             // jog to position
             //*********************************************************************************************************
           ELSIF #tempJogToPosition THEN
             // set jog target position and configuration
             #instMC_MoveLinearAbsoute.Position[1] := #targetPosition.x;
             #instMC_MoveLinearAbsoute.Position[2] := #targetPosition.y;
             #instMC_MoveLinearAbsoute.Position[3] := #targetPosition.z;
             #instMC_MoveLinearAbsoute.Position[4] := #targetPosition.a;
             #instMC_MoveLinearAbsoute.CoordSystem := #coordSystem;
             #instMC_MoveLinearAbsoute.Velocity := #dynamics.path.velocity;
             #instMC_MoveLinearAbsoute.Acceleration := #dynamics.path.acceleration;
             #instMC_MoveLinearAbsoute.Deceleration := #dynamics.path.deceleration;
             #instMC_MoveLinearAbsoute.Jerk := #dynamics.path.jerk;
             #instMC_MoveLinearAbsoute.DynamicAdaption := #dynamics.dynamicAdaption;
           END_IF;

         END_REGION

         REGION STATE_TRANSITION

           // check if change of tool is required
           IF (#tool <> #statToolOld) THEN
             #statFBState := #FB_STATE_SET_TOOL;

             // check if orientation movement required
           ELSIF (((#jogDirection = 4) AND (#tempJogForward OR #tempJogBackward)) OR #tempJogToPosition)
             AND (#dynamics.orientation.velocity > 0.0 // check if change of orientation dynamics is required
             OR #dynamics.orientation.acceleration > 0.0
             OR #dynamics.orientation.deceleration > 0.0
             OR #dynamics.orientation.jerk > 0.0)
           THEN
             #statFBState := #FB_STATE_SET_DYNAMICS;

             // execute movement
           ELSE
             #statFBState := #FB_STATE_EXECUTE_MOVEMENT;
           END_IF;

         END_REGION

       #FB_STATE_SET_TOOL:

         REGION TOOL_CHANGE

           IF #axesGroup.StatusWord.%X6 // no motion command is acitve
             AND NOT #axesGroup.StatusWord.%X17 // not interrupted
             AND #axesGroup.StatusWord.%X12 // constant velocity
           THEN
             #instMC_SetTool.Execute := TRUE;
             #instMC_SetTool.ToolNumber := #tool;
           END_IF;

         END_REGION

         REGION STATE_TRANSITION

           // tool has been changed
           IF #instMC_SetTool.Done THEN
             #statToolOld := #tool;

             // check if orientation movement required
             IF (((#jogDirection = 4) AND (#tempJogForward OR #tempJogBackward)) OR #tempJogToPosition)
               AND (#dynamics.orientation.velocity > 0.0 // check if change of orientation dynamics is required
               OR #dynamics.orientation.acceleration > 0.0
               OR #dynamics.orientation.deceleration > 0.0
               OR #dynamics.orientation.jerk > 0.0)
             THEN
               #statFBState := #FB_STATE_SET_DYNAMICS;

               // execute movement  
             ELSE
               #statFBState := #FB_STATE_EXECUTE_MOVEMENT;
             END_IF;
           END_IF;

         END_REGION

       #FB_STATE_SET_DYNAMICS:

         REGION SET_ORIENTATION_DYNAMICS

           // safe default dynimcs for orientation axis
           #statOrientationDynamicsOld.velocity := #axesGroup.DynamicDefaults.Orientation.Velocity;
           #statOrientationDynamicsOld.acceleration := #axesGroup.DynamicDefaults.Orientation.Acceleration;
           #statOrientationDynamicsOld.deceleration := #axesGroup.DynamicDefaults.Orientation.Deceleration;
           #statOrientationDynamicsOld.jerk := #axesGroup.DynamicDefaults.Orientation.Jerk;

           // change orientation default dynamics temporary
           #axesGroup.DynamicDefaults.Orientation.Velocity := #dynamics.orientation.velocity;
           #axesGroup.DynamicDefaults.Orientation.Acceleration := #dynamics.orientation.acceleration;
           #axesGroup.DynamicDefaults.Orientation.Deceleration := #dynamics.orientation.deceleration;
           #axesGroup.DynamicDefaults.Orientation.Jerk := #dynamics.orientation.jerk;

           // Orientation default dynamics will be reseted to previous values after jogging
           #statOrientationDynamicsChanged := TRUE;

         END_REGION

         // FB state transition 
         #statFBState := #FB_STATE_EXECUTE_MOVEMENT;

       #FB_STATE_EXECUTE_MOVEMENT:

         REGION SET_JOG_COMMAND

           // Cartesian jogging
           IF (#tempJogForward OR #tempJogBackward) THEN
             #instMC_MoveLinearRelative.Execute := TRUE;

             // jog to target position  
           ELSIF #tempJogToPosition THEN
             #instMC_MoveLinearAbsoute.Execute := TRUE;
           ELSE
             #instMC_MoveLinearRelative.Execute := FALSE;
             #instMC_MoveLinearAbsoute.Execute := FALSE;
           END_IF;

         END_REGION

         REGION STATE_TRANSITION

           IF #instMC_MoveLinearRelative.Done OR #instMC_MoveLinearAbsoute.Done THEN
             #statStatus := #STATUS_EXECUTION_FINISHED;
           END_IF;

         END_REGION

       #FB_STATE_STOP:

         REGION STOP_KINEMATICS_MOTION

           // set execute if group stop not busy
           IF NOT #instMC_GroupStop.Busy AND NOT #instMC_GroupStop.Done AND NOT #instMC_GroupStop.Error THEN
             #instMC_GroupStop.Execute := TRUE;
           ELSE
             #instMC_GroupStop.Execute := FALSE;
           END_IF;

         END_REGION

         REGION STATE_TRANSITION

           IF #instMC_GroupStop.Done THEN
             #statStatus := #STATUS_EXECUTION_FINISHED;
           ELSIF #axesGroup.StatusWord.%X1 THEN // general TO error
             #statStatus := #ERR_TO_KINEMATICS;
           ELSIF #instMC_MoveLinearRelative.Error THEN
             #statStatus := #instMC_MoveLinearRelative.ErrorId;
           ELSIF #instMC_MoveLinearAbsoute.Error THEN
             #statStatus := #instMC_MoveLinearAbsoute.ErrorId;
           ELSIF #instMC_SetTool.Error THEN
             #statStatus := #instMC_SetTool.ErrorId;
           ELSIF #instMC_GroupStop.Error THEN
             #statStatus := #instMC_GroupStop.ErrorId;
           END_IF;

         END_REGION

       ELSE // Undefined state in state machine reached
         #statStatus := #ERR_UNDEFINED_STATE;
     END_CASE;

   END_REGION STATE_MACHINE

   REGION OUTPUTS

     // Write outputs
     IF (#statStatus = #STATUS_EXECUTION_FINISHED) AND (#statDone = FALSE) AND (#statError = FALSE) THEN // Execution finished without errors
       #statDone := TRUE;
       #statBusy := FALSE;
       #statActive := FALSE;
       #statError := FALSE;
       #statFBState := #FB_STATE_NO_PROCESSING; // Switch state machine to "no processing"

     ELSIF (#statStatus.%X15 = TRUE) AND (#statError = FALSE) THEN // Error occurred (#statStatus is 16#8000 to 16#FFFF)
       #statDone := FALSE;
       #statBusy := FALSE;
       #statActive := FALSE;
       #statError := TRUE;
       // Write diagnostics
       #tempRet := RD_SYS_T(#diagnostics.timeStamp);
       #diagnostics.stateNumber := #statFBState;
       #diagnostics.status := #statStatus;
       #statFBState := #FB_STATE_NO_PROCESSING; // Switch state machine to "no processing"

     ELSIF (#tempJogForward = FALSE AND #tempJogBackward = FALSE AND #tempJogToPosition = FALSE) AND ((#statDone = TRUE) OR (#statError = TRUE)) THEN // Reset outputs
       #statDone := FALSE;
       #statBusy := FALSE;
       #statActive := FALSE;
       #statError := FALSE;
       #statStatus := #STATUS_NO_CALL;
       #statJogForwardOld := FALSE;
       #statJogBackwardOld := FALSE;
       #statJogToPositionOld := FALSE;
     END_IF;

     // Write static values to outputs
     #done := #statDone;
     #busy := #statBusy;
     #active := #statActive;
     #error := #statError;
     #status := #statStatus;
     #remainingDistance := #statRemainingDistance;

   END_REGION OUTPUTS

   REGION CALL_FB_CYCLICALLY

     // call FBs and set Execute = FALSE after the call
     #instMC_GroupStop(AxesGroup := #axesGroup);
     #instMC_GroupStop.Execute := FALSE;

     #instMC_MoveLinearAbsoute(AxesGroup := #axesGroup);
     #instMC_MoveLinearAbsoute.Execute := FALSE;

     #instMC_MoveLinearRelative(AxesGroup := #axesGroup);
     #instMC_MoveLinearRelative.Execute := FALSE;

     #instMC_SetTool(AxesGroup := #axesGroup);
     #instMC_SetTool.Execute := FALSE;

   END_REGION
END_FUNCTION_BLOCK

FUNCTION "LKinCtrl_MC_PathSelect" : "LKinCtrl_typeDiagnosticsPathSelect"   // FC35001, SCL
TITLE = LKinCtrl_MC_PathSelect
{ S7_Optimized_Access := 'TRUE' }
AUTHOR : tech.team.motioncontrol@siemens.com
FAMILY : LKinCtrl
VERSION : 1.0
// The FC creates a command list (PathData) for execution with FB LKinCtrl_MovePath.
   VAR_IN_OUT
      pathDescription : "LKinCtrl_typePathDescription";   // point table containing path points
      pathData : Variant;   // generated PathData from point table
   END_VAR
   VAR_TEMP
      tempPathData_reduced : REF_TO "LKinCtrl_typePathData_reduced";   // temporary reference to PathData_reduced
      tempPathData_advanced : REF_TO "LKinCtrl_typePathData_advanced";   // temporary reference to PathData_advanced
      tempPathData : REF_TO "LKinCtrl_typePathData";   // temporary reference to PathData
      tempPathDataType : Int;   // temporary variable storing detected PathData type
      tempPointLimit : Int;   // temporary variable storing end of point array
      tempPathDataLimit : Int;   // temporary variable storing end of pathData
      tempCtr : Int;   // temporary counter
      tempFlagCtr : Int;   // temporary flag counter
      tempPathDataElementCtr : Int;   // temporary path data element counter
      tempPathDataElement : "LKinCtrl_typePathDataElement";   // temporary path data element
      tempPointEmpty : "LKinCtrl_typePathDescriptionElement";   // temporary empty path description element
      tempEmptyFlag : "LKinCtrl_typeSetFlagElement_Bool";   // temporary empty flag element
      tempEmptyValueFlag : "LKinCtrl_typeSetFlagElement_LReal";   // temporary empty value flag element
   END_VAR
   // Ret_Val : return value struct of this function
   VAR CONSTANT
      STATUS_EXECUTION_FINISHED : Word := 16#0000;   // status PathData generated without error
      ERR_WRONG_CS : Word := 16#8280;   // error due to an incorrect defined CS
      ERR_WRONG_FLAG : Word := 16#8281;   // error due to an incorrect flag definition
      ERR_WRONG_FLAGMODE : Word := 16#8282;   // error due to an incorrect flagMode definition
      ERR_PATHDATA_OVERFLOW : Word := 16#8283;   // error due to more points than path data elements
      ERR_UNDEFINED_STATE : Word := 16#8600;   // error due to an undefined FB state
   END_VAR
BEGIN
   //==========================================================================================
   // SIEMENS AG
   // (c)Copyright 2020 All Rights Reserved
   //------------------------------------------------------------------------------------------
   // Library: LKinCtrl
   // Tested with: S7-1517T-3 PN/DP
   // Engineering: TIA Portal V15
   // Restrictions: ---
   // Requirements: S7-1500T FW 2.5
   // Functionality: MC_PathSelect
   // The FC creates a command list (PathData) for execution with FB LKinCtrl_MovePath.
   // The data for the creation of the path provided by a point list (PathDescription)
   // 
   // Support: tech.team.motioncontrol@siemens.com
   // Note: Parameter comments are only available in language 'English (United States)'
   //------------------------------------------------------------------------------------------
   // Change log table:
   // Version    Date          Expert in charge    Changes applied
   // 01.00.00   01.04.2018    JR / FR             First release version v1.0,
   // 01.00.01   30.01.2020    FR                  Removed commented code & changed flag constant
   // 01.00.02   13.02.2020    FR                  Initialize emptyPoint flag structure correctly
   // 01.00.03   18.03.2020    FR                  Added valueFlags to point
   //===========================================================================================
   // Initialize return value
   #LKinCtrl_MC_PathSelect.#status := #ERR_UNDEFINED_STATE;

   // Initialize pathdata counter
   #tempPathDataElementCtr := 1;

   // Initialize pathDesription limit
   #tempPointLimit := "LKINCTRL_NO_OF_PATHDATA_ELEMENTS";

   // Initialize emptyPoint flag structure
   FOR #tempCtr := 1 TO "LKINCTRL_NO_OF_CMD_SETFLAGS" DO
     #tempPointEmpty.flags[#tempCtr] := #tempEmptyFlag;
   END_FOR;

   // Initialize emptyPoint valueFlag structure
   FOR #tempCtr := 1 TO "LKINCTRL_NO_OF_CMD_VALUEFLAGS" DO
     #tempPointEmpty.valueFlags[#tempCtr] := #tempEmptyValueFlag;
   END_FOR;

   REGION PATHDATA_CONVERSION
     // reduced PathData (only linear commands with blending and dynamics)
     IF TypeOf(#pathData) = LKinCtrl_typePathData_reduced THEN
       #tempPathData_reduced ?= #pathData;
       #tempPathDataType := "LKINCTRL_PATHDATA_TYPE_REDUCED";
       #tempPathDataLimit := "LKINCTRL_NO_OF_PATHDATA_ELEMENTS_REDUCED";

       // regular PathData (no pointers)
     ELSIF TypeOf(#pathData) = LKinCtrl_typePathData THEN
       #tempPathData ?= #pathData;
       #tempPathDataType := "LKINCTRL_PATHDATA_TYPE_NORMAL";
       #tempPathDataLimit := "LKINCTRL_NO_OF_PATHDATA_ELEMENTS";

       // advanced PathData (all elements)
     ELSIF TypeOf(#pathData) = LKinCtrl_typePathData_advanced THEN
       #tempPathData_advanced ?= #pathData;
       #tempPathDataType := "LKINCTRL_PATHDATA_TYPE_ADVANCED";
       #tempPathDataLimit := "LKINCTRL_NO_OF_PATHDATA_ELEMENTS_ADVANCED";
     END_IF;
   END_REGION PATHDATA_CONVERSION 

   // For loop over all elements in path data
   FOR #tempCtr := 1 TO #tempPointLimit DO
     // Check path data length
     IF #tempCtr <= #tempPathDataLimit THEN

         // CHECK FOR COMMAND TO BE ACTIVE / SET IN POINT TABLE
         IF #pathDescription.points[#tempCtr] = #tempPointEmpty THEN
           ; // done
           #LKinCtrl_MC_PathSelect.status := #STATUS_EXECUTION_FINISHED;
           RETURN;
         ELSE
           // Copy command
           REGION COPY_TO_TEMP
             #tempPathDataElement.cmdType := 1;
             #tempPathDataElement.cmdName := #pathDescription.points[#tempCtr].pointName;
             #tempPathDataElement.cmdCoordinates.cartesianPosition := #pathDescription.points[#tempCtr].targetPosition;

             // Check CoordSystem 
             IF #pathDescription.points[#tempCtr].coordSystem > -1
               AND #pathDescription.points[#tempCtr].coordSystem < 4
             THEN
               #tempPathDataElement.cmdCoordinates.coordSystem := #pathDescription.points[#tempCtr].coordSystem;
             ELSE
               // error handling
               #LKinCtrl_MC_PathSelect.status := #ERR_WRONG_CS;
               #LKinCtrl_MC_PathSelect.entryID := #tempCtr;
               RETURN;
             END_IF;

             // Copy blending radius
             #tempPathDataElement.cmdParameters.transitionParameters[1] := #pathDescription.points[#tempCtr].blendingDistance;

             // Check bufferMode
             IF #pathDescription.points[#tempCtr].blendingDistance <> 0.0 THEN
               // set bufferMode to BM_BLENDING_HIGH by default if blending distance <> 0.0
               #tempPathDataElement.cmdParameters.bufferMode := 5;
             ELSE
               // set bufferMode to BM_BUFFERD by default if blending distance = 0.0
               #tempPathDataElement.cmdParameters.bufferMode := 1;
             END_IF;

             // Check setFlags
             FOR #tempFlagCtr := 1 TO "LKINCTRL_NO_OF_CMD_SETFLAGS" DO
               // check flag number to be valid
               IF #pathDescription.points[#tempCtr].flags[#tempFlagCtr].flag >= -1
                 AND #pathDescription.points[#tempCtr].flags[#tempFlagCtr].flag <= "LKINCTRL_NO_OF_LAST_SETFLAG"
               THEN
                 #tempPathDataElement.setFlags[#tempFlagCtr].flag := #pathDescription.points[#tempCtr].flags[#tempFlagCtr].flag;
               ELSE
                 // error handling
                 #LKinCtrl_MC_PathSelect.status := #ERR_WRONG_FLAG;
                 #LKinCtrl_MC_PathSelect.entryID := #tempCtr;
                 RETURN;
               END_IF;

               // check flagmode to be valid
               IF #pathDescription.points[#tempCtr].flags[#tempFlagCtr].flagMode = 0
                 OR #pathDescription.points[#tempCtr].flags[#tempFlagCtr].flagMode = 1
                 OR #pathDescription.points[#tempCtr].flags[#tempFlagCtr].flagMode = 2
                 OR #pathDescription.points[#tempCtr].flags[#tempFlagCtr].flagMode = 3
                 OR #pathDescription.points[#tempCtr].flags[#tempFlagCtr].flagMode = 5
                 OR #pathDescription.points[#tempCtr].flags[#tempFlagCtr].flagMode = 10
                 OR #pathDescription.points[#tempCtr].flags[#tempFlagCtr].flagMode = 11
                 OR #pathDescription.points[#tempCtr].flags[#tempFlagCtr].flagMode = 13
               THEN
                 #tempPathDataElement.setFlags[#tempFlagCtr].flagMode := #pathDescription.points[#tempCtr].flags[#tempFlagCtr].flagMode;
               ELSE
                 // error handling
                 #LKinCtrl_MC_PathSelect.status := #ERR_WRONG_FLAGMODE;
                 #LKinCtrl_MC_PathSelect.entryID := #tempCtr;
                 RETURN;
               END_IF;
             END_FOR;

             // Check valueFlags
             FOR #tempFlagCtr := 1 TO "LKINCTRL_NO_OF_CMD_VALUEFLAGS" DO
               // check flag number to be valid
               IF #pathDescription.points[#tempCtr].valueFlags[#tempFlagCtr].flag >= -1
                 AND #pathDescription.points[#tempCtr].valueFlags[#tempFlagCtr].flag <= "LKINCTRL_NO_OF_LAST_VALUEFLAG"
               THEN
                 // Set flag number
                 #tempPathDataElement.valueFlags[#tempFlagCtr].flag := #pathDescription.points[#tempCtr].valueFlags[#tempFlagCtr].flag;
               ELSE
                 // error handling
                 #LKinCtrl_MC_PathSelect.status := #ERR_WRONG_FLAG;
                 #LKinCtrl_MC_PathSelect.entryID := #tempCtr;
                 RETURN;
               END_IF;

               // check flagmode to be valid
               IF #pathDescription.points[#tempCtr].valueFlags[#tempFlagCtr].flagMode = 0
                 OR #pathDescription.points[#tempCtr].valueFlags[#tempFlagCtr].flagMode = 1
                 OR #pathDescription.points[#tempCtr].valueFlags[#tempFlagCtr].flagMode = 2
                 OR #pathDescription.points[#tempCtr].valueFlags[#tempFlagCtr].flagMode = 3
                 OR #pathDescription.points[#tempCtr].valueFlags[#tempFlagCtr].flagMode = 5
                 OR #pathDescription.points[#tempCtr].valueFlags[#tempFlagCtr].flagMode = 10
                 OR #pathDescription.points[#tempCtr].valueFlags[#tempFlagCtr].flagMode = 11
                 OR #pathDescription.points[#tempCtr].valueFlags[#tempFlagCtr].flagMode = 13
               THEN
                 // Set flagMode and Value
                 #tempPathDataElement.valueFlags[#tempFlagCtr].flagMode := #pathDescription.points[#tempCtr].valueFlags[#tempFlagCtr].flagMode;
                 #tempPathDataElement.valueFlags[#tempFlagCtr].value := #pathDescription.points[#tempCtr].valueFlags[#tempFlagCtr].value;
               ELSE
                 // error handling
                 #LKinCtrl_MC_PathSelect.status := #ERR_WRONG_FLAGMODE;
                 #LKinCtrl_MC_PathSelect.entryID := #tempCtr;
                 RETURN;
               END_IF;
             END_FOR;
           END_REGION COPY_TO_TEMP

           REGION COPY_TO_OUTPUT
             CASE #tempPathDataType OF
               "LKINCTRL_PATHDATA_TYPE_REDUCED": // Path data reduced
                 // Copy command
                 #tempPathData_reduced<?OpDeref?>.commands[#tempPathDataElementCtr].cmdType := #tempPathDataElement.cmdType;
                 #tempPathData_reduced<?OpDeref?>.commands[#tempPathDataElementCtr].cmdName := #tempPathDataElement.cmdName;
                 #tempPathData_reduced<?OpDeref?>.commands[#tempPathDataElementCtr].cmdActivated := #tempPathDataElement.cmdActivated; // !
                 #tempPathData_reduced<?OpDeref?>.commands[#tempPathDataElementCtr].cmdCoordinates := #tempPathDataElement.cmdCoordinates;
                 #tempPathData_reduced<?OpDeref?>.commands[#tempPathDataElementCtr].cmdParameters.bufferMode := #tempPathDataElement.cmdParameters.bufferMode;
                 #tempPathData_reduced<?OpDeref?>.commands[#tempPathDataElementCtr].cmdParameters.transitionParameters[1] := #tempPathDataElement.cmdParameters.transitionParameters[1];
                 #tempPathData_reduced<?OpDeref?>.commands[#tempPathDataElementCtr].setFlags := #tempPathDataElement.setFlags;
                 #tempPathData_reduced<?OpDeref?>.commands[#tempPathDataElementCtr].valueFlags := #tempPathDataElement.valueFlags;

               "LKINCTRL_PATHDATA_TYPE_NORMAL": // Path data normal
                 #tempPathData<?OpDeref?>.commands[#tempPathDataElementCtr] := #tempPathDataElement;

               "LKINCTRL_PATHDATA_TYPE_ADVANCED": // Path data advanced
                 // Copy command
                 #tempPathData_advanced<?OpDeref?>.commands[#tempPathDataElementCtr].cmdType := #tempPathDataElement.cmdType;
                 #tempPathData_advanced<?OpDeref?>.commands[#tempPathDataElementCtr].cmdName := #tempPathDataElement.cmdName;
                 #tempPathData_advanced<?OpDeref?>.commands[#tempPathDataElementCtr].cmdActivated := #tempPathDataElement.cmdActivated; // !
                 #tempPathData_advanced<?OpDeref?>.commands[#tempPathDataElementCtr].cmdCoordinates := #tempPathDataElement.cmdCoordinates;
                 #tempPathData_advanced<?OpDeref?>.commands[#tempPathDataElementCtr].cmdParameters := #tempPathDataElement.cmdParameters;
                 #tempPathData_advanced<?OpDeref?>.commands[#tempPathDataElementCtr].setFlags := #tempPathDataElement.setFlags;
                 #tempPathData_advanced<?OpDeref?>.commands[#tempPathDataElementCtr].valueFlags := #tempPathDataElement.valueFlags;

               ELSE  // Wrong pathData type?
                 #LKinCtrl_MC_PathSelect.#status := #ERR_UNDEFINED_STATE;
             END_CASE;

             // Increment counter for path data element
             #tempPathDataElementCtr += 1;

           END_REGION COPY_TO_OUTPUT
       END_IF;

     ELSE
       // Error more points than path data elements
       #LKinCtrl_MC_PathSelect.status := #ERR_PATHDATA_OVERFLOW;
       #LKinCtrl_MC_PathSelect.entryID := #tempCtr;
       RETURN;
     END_IF;
   END_FOR;

   // Write return value 
   #LKinCtrl_MC_PathSelect.status := #STATUS_EXECUTION_FINISHED;

   // =================================================================================================================
   // End of Function: LKinCtrl_MC_PathSelect
   // =================================================================================================================
END_FUNCTION

// folder: LKinCtrl_Blocks/LKinCtrl_AuxBlocks

FUNCTION_BLOCK "LKinCtrl_GetKinematicsStatusWord"   // FB35004, SCL
TITLE = LKinCtrl_GetKinematicsStatusWord
{ S7_Optimized_Access := 'TRUE' }
AUTHOR : tech.team.motioncontrol@siemens.com
FAMILY : LKinCtrl
VERSION : 1.0
// FB provides functionalities to reveice status information on Kinematics StatusWord
   VAR_INPUT
      axesGroup : TO_Kinematics;   // reference to the axesGroup
   END_VAR
   VAR_OUTPUT
      error : Bool;   // error axesGroup
      restartActive : Bool;   // restart of TO Kinematic active
      onlineStartValuesChanged : Bool;   // change of start values TO Kinematic
      controlPanelActive : Bool;   // control panel TO Kinematic activated
      done : Bool;   // no motion command active / control panel deactivated
      linearCommand : Bool;   // linear command active
      circularCommand : Bool;   // circular command active
      constantVelocity : Bool;   // TO Kinematic at constant velocity
      accelerating : Bool;   // acceleration progress active
      decelerating : Bool;   // deceleration progress active
      orientationMotion : Bool;   // orientation motion active
      stopping : Bool;   // MC_GroupStop is active
      interrupted : Bool;   // motion interrupted
      blending : Bool;   // no blending segment active
   END_VAR
   VAR
      statFirstCycle : Bool := TRUE;   // flag first cycle
      statStatusWordOld : DWord;   // flag word for old statusWord
   END_VAR
   VAR_TEMP
      tempStatusWord : DWord;
   END_VAR
BEGIN
   //==========================================================================================
   // SIEMENS AG
   // (c)Copyright 2019 All Rights Reserved
   //------------------------------------------------------------------------------------------
   // Library: LKinCtrl
   // Tested with: S7-1515T-2 PN
   // Engineering: TIA Portal V15
   // Restrictions: ---
   // Requirements: S7-1500T FW 2.5
   // Functionality: LKinCtrl_GetKinematicsStatusWord
   // The FB is splitting the status word of a technoloy object kinematic into bits.
   // Support: tech.team.motioncontrol@siemens.com
   // Note: Parameter comments are only available in language 'English (United States)'
   //------------------------------------------------------------------------------------------
   // Change log table:
   // Version    Date          Expert in charge    Changes applied
   // 01.00.00   16.08.2017    RK                  First released version
   //===========================================================================================

   //----------------------------------------------------------------------------------------------
   // Read statusword
   //----------------------------------------------------------------------------------------------
   #tempStatusWord := #axesGroup.StatusWord;

   //----------------------------------------------------------------------------------------------
   // Write outputs
   //----------------------------------------------------------------------------------------------
   IF #tempStatusWord <> #statStatusWordOld
       OR #statFirstCycle
   THEN
       #error := #tempStatusWord.%X1;
       #restartActive := #tempStatusWord.%X2;
       #onlineStartValuesChanged := #tempStatusWord.%X3;
       #controlPanelActive := #tempStatusWord.%X4;
       // #reservedBit_5 := #tempStatusWord.%X5;
       #done := #tempStatusWord.%X6;
       // #reservedBit_7 := #tempStatusWord.%X7;
       #linearCommand := #tempStatusWord.%X8;
       #circularCommand := #tempStatusWord.%X9;
       // #polynomialCommand := #tempStatusWord.%X10;
       // #directCommand := #tempStatusWord.%X11;
       #constantVelocity := #tempStatusWord.%X12;
       #accelerating := #tempStatusWord.%X13;
       #decelerating := #tempStatusWord.%X14;
       #orientationMotion := #tempStatusWord.%X15;
       #stopping := #tempStatusWord.%X16;
       #interrupted := #tempStatusWord.%X17;
       #blending := #tempStatusWord.%X18;

       // Set back flag
       #statFirstCycle := False;
   ELSE
       ; // Do nothing
   END_IF;

   // Copy current state of status for edge detection
   #statStatusWordOld := #tempStatusWord;
END_FUNCTION_BLOCK

FUNCTION_BLOCK "LKinCtrl_GetKinematicsErrorWord"   // FB35005, SCL
TITLE = LKinCtrl_GetKinematicsErrorWord
{ S7_Optimized_Access := 'TRUE' }
AUTHOR : tech.team.motioncontrol@siemens.com
FAMILY : LKinCtrl
VERSION : 1.0
// FB provides functionalities to reveice status information on Kinematics ErrorWord
   VAR_INPUT
      axesGroup : TO_Kinematics;   // reference to the axesGroup
   END_VAR
   VAR_OUTPUT
      systemFault : Bool;   // system-internal error has occured
      configFault : Bool;   // one or more configuration parameters are inconsistent or invalid
      userFault : Bool;   // error in the user program with a Motion Control instructioc or its use
      commandNotAccepted : Bool;   // command cannot be accepted
      transformationFault : Bool;   // error in the kinematics transformation
      dynamicError : Bool;   // specified dynamic values are limited to permissible values
   END_VAR
   VAR
      statFirstCycle : Bool := TRUE;   // flag first cycle
      statErrorWordOld : DWord;   // flag word for old errorWord
   END_VAR
   VAR_TEMP
      tempErrorWord : DWord;
   END_VAR
BEGIN
   //==========================================================================================
   // SIEMENS AG
   // (c)Copyright 2019 All Rights Reserved
   //------------------------------------------------------------------------------------------
   // Library: LKinCtrl
   // Tested with: S7-1515T-2 PN
   // Engineering: TIA Portal V15
   // Restrictions: ---
   // Requirements: S7-1500T FW 2.5
   // Functionality: LKinCtrl_GetKinematicsErrorWord
   // The FB is splitting the error word of a technoloy object kinematic into bits.
   // Support: tech.team.motioncontrol@siemens.com
   // Note: Parameter comments are only available in language 'English (United States)'
   //------------------------------------------------------------------------------------------
   // Change log table:
   // Version    Date          Expert in charge    Changes applied
   // 01.00.00   16.08.2017    RK                  First released version
   //===========================================================================================

   //----------------------------------------------------------------------------------------------
   // Read errorWord
   //----------------------------------------------------------------------------------------------
   #tempErrorWord := #axesGroup.ErrorWord;

   //----------------------------------------------------------------------------------------------
   // Write outputs
   //----------------------------------------------------------------------------------------------
   IF #tempErrorWord <> #statErrorWordOld
       OR #statFirstCycle
     THEN
       #systemFault := #tempErrorWord.%X0;
       #configFault := #tempErrorWord.%X1;
       #userFault := #tempErrorWord.%X2;
       #commandNotAccepted := #tempErrorWord.%X3;
       #transformationFault := #tempErrorWord.%X4;
       #dynamicError := #tempErrorWord.%X6;


       // Set back flag
       #statFirstCycle := False;
   ELSE
       ; // Do nothing
   END_IF;

   // Copy current state of error for edge detection
   #statErrorWordOld := #tempErrorWord;
END_FUNCTION_BLOCK

FUNCTION_BLOCK "LKinCtrl_GetKinematicsWarningWord"   // FB35006, SCL
TITLE = LKinCtrl_GetKinematicsWarningWord
{ S7_Optimized_Access := 'TRUE' }
AUTHOR : tech.team.motioncontrol@siemens.com
FAMILY : LKinCtrl
VERSION : 1.0
// FB provides functionalities to reveice status information on Kinematics WarningWord
   VAR_INPUT
      axesGroup : TO_Kinematics;   // reference to the axesGroup
   END_VAR
   VAR_OUTPUT
      systemFault : Bool;   // system-internal error has occured
      configFault : Bool;   // one or more configuration parameters are inconsistent or invalid
      userFault : Bool;   // error in the user program with a Motion Control instructioc or its use
      commandNotAccepted : Bool;   // command cannot be accepted
      dynamicWarning : Bool;   // specified dynamic values are limited to permissible values
   END_VAR
   VAR
      statFirstCycle : Bool := TRUE;   // flag first cycle
      statWarningWordOld : DWord;   // flag word for old warningWord
   END_VAR
   VAR_TEMP
      tempWarningWord : DWord;
   END_VAR
BEGIN
   //==========================================================================================
   // SIEMENS AG
   // (c)Copyright 2019 All Rights Reserved
   //------------------------------------------------------------------------------------------
   // Library: LKinCtrl
   // Tested with: S7-1515T-2 PN
   // Engineering: TIA Portal V15
   // Restrictions: ---
   // Requirements: S7-1500T FW 2.5
   // Functionality: LinCtrl_GetKinematicsWarningWord
   // The FB is splitting the warning word of a technoloy object kinematic into bits.
   // Support: tech.team.motioncontrol@siemens.com
   // Note: Parameter comments are only available in language 'English (United States)'
   //------------------------------------------------------------------------------------------
   // Change log table:
   // Version    Date          Expert in charge    Changes applied
   // 01.00.00   16.08.2017    RK                  First released version
   //===========================================================================================

   //----------------------------------------------------------------------------------------------
   // Read warningWord
   //----------------------------------------------------------------------------------------------
   #tempWarningWord := #axesGroup.WarningWord;

   //-----------------------------------------------
   //
   //
   //-----------------------------------------------
   // Write outputs
   //----------------------------------------------------------------------------------------------
   IF #tempWarningWord <> #statWarningWordOld
       OR #statFirstCycle
     THEN
       #systemFault := #tempWarningWord.%X0;
       #configFault := #tempWarningWord.%X1;
       #userFault := #tempWarningWord.%X2;
       #commandNotAccepted := #tempWarningWord.%X3;
       #dynamicWarning := #tempWarningWord.%X6;


       // Set back flag
       #statFirstCycle := False;
   ELSE
       ; // Do nothing
   END_IF;

   // Copy current state of warning for edge detection
   #statWarningWordOld := #tempWarningWord;
END_FUNCTION_BLOCK

FUNCTION_BLOCK "LKinCtrl_MC_GroupPower"   // FB35021, SCL
TITLE = LKinCtrl_MC_GroupPower
{ S7_Optimized_Access := 'TRUE' }
AUTHOR : tech.team.motioncontrol@siemens.com
FAMILY : LKinCtrl
VERSION : 2.0
// FB provides funcitonalities to enable all axes (TO_PositioningAxis or TO_SynchronousAxis) interconnected with TO Kinematics
   VAR_INPUT
      enable : Bool;   // TRUE: Enable axes; FALSE: Disable axes
      startMode : Array[1..#MAX_NO_OF_AXES] of DInt;   // startMode of axis; 0: enable NOT position controlled; 1: enable position controlled
      stopMode : Array[1..#MAX_NO_OF_AXES] of Int;   // stopMode of axis; 0: emergency stop; 1: immediate stop; 2: stop with max dynamics
   END_VAR
   VAR_OUTPUT
      busy : Bool;   // TRUE: FB is not finished and new output values can be expected
      error : Bool;   // TRUE: An error occurred during the execution of the FB
      axesEnabled : Bool := false;   // TRUE: all axes of axesGroup enabled; FALSE: all axes of axesGroup disabled
      diagnostics : "LKinCtrl_typeAuxFCDiagnostics";   // Diagnostics information of FB (optional)
   END_VAR
   VAR_IN_OUT
      axesGroup : TO_Kinematics;   // reference to the axesGroup
   END_VAR
   VAR
      statEnableOld : Bool;   // old value of 'enable' input for edge detection
      statBusy : Bool;   // static value for output 'busy'
      statError : Bool;   // static value for output 'error'
      statErrorUserCleared : Bool;   // error occurred that can only be solved by user; rising edge at enable input necessary
      statErrorAutoCleared : Bool;   // error occurred that can be acknowledged by FB
      statStatus : Word := 16#7000;   // static value for output 'status'
      statSubfunctionStatus : Word;   // static value for output 'subFunctionStatus'
      statAxesEnabled : Bool;   // static value for output 'axesEnabled'
      statAxesDisabled : Bool;   // static value for output 'axesDisabled'
      statErrorDetailNumber : UDInt;   // static to store axis error detail number
      statStateMachine : DInt := 0;   // state in the state machine of the FB
      statDisablingCompleted : Bool;   // TRUE: Disabling has been completed
      statAxisNumberDiag : Int;   // static value for output 'axisNumber'
      instMC_Power : Array[1..#MAX_NO_OF_AXES] of MC_POWER;   // multi instance array of MC_RESET for axes
      statEnableAxis : Array[1..#MAX_NO_OF_AXES] of Bool;   // array of execute triggers for MC_HOME
      statAxes : Array[1..#MAX_NO_OF_AXES] of Struct   // array of struct containing axis DB_ANY and type of axis
         typeOfAxis : Int;
         axis : DB_ANY;
      END_STRUCT;
      statAxisStatusWord : DWord;   // static to store axis status word
      statAxisErrorDetailNumber : UDInt;   // static to store axis error detail number
      statExsitingAxesCtr : Int;   // static counter for existing axes
      statEnabledAxesCtr : Int;   // static counter for enabled axes
      statDisabledAxesCtr : Int;   // static counter for disabled axes
   END_VAR
   VAR_TEMP
      tempEnable : Bool;   // temporary value for input 'enable'
      tempAxisCtr : Int;   // temporary counter variable for axes
   END_VAR
   VAR CONSTANT
      NO_PROCESSING : DInt := 0;   // FB state: No processing
      DETECT_AXES : DInt := 10;   // state machine constant
      CHECK_AXES : DInt := 40;   // state machine constant
      ENABLING_AXES : DInt := 50;   // state machine constant
      ENABLED_AXES : DInt := 55;   // state machine constant
      DISABLING_AXES : DInt := 60;   // state machine constant
      DISABLED_AXES : DInt := 65;   // state machine constant
      AXIS_NOT_USED : Int := -1;   // type of axis constant
      TYPE_POSITIONING_AXIS : Int := 0;   // type of axis constant
      TYPE_SYNCHRONOUS_AXIS : Int := 1;   // type of axis constant
      MAX_NO_OF_AXES : Int := 4;   // maximum number of axes
      ERROR_STATE : DInt := 90;   // state machine constant
      STATUS_NO_ERROR : Word := 16#0000;   // no error occured
      STATUS_NO_CALL : Word := 16#7000;   // no job being currently processed
      STATUS_FIRST_CALL : Word := 16#7001;   // first call after incoming new job (rising edge 'execute')
      STATUS_SUBSEQUENT_CALL : Word := 16#7002;   // subsequent call during active processing without further details
      STATUS_ENABLING_AXES_IN_PROGRESS : Word := 16#7008;   // enabling axes in progress
      STATUS_DISABLING_AXES_IN_PROGRESS : Word := 16#7010;   // disabling axes in progress
      STATUS_ALL_AXES_ENABLED : Word := 16#7009;   // all access enabled successfully
      STATUS_ALL_AXES_DISABLED : Word := 16#7011;   // all access disabled successfully
      ERR_UNDEFINED_STATE : Word := 16#8600;   // error due to an undefined state in state machine
      ERR_AXIS_ERROR : Word := 16#8370;   // error pending at axis
      ERR_KIN_ERROR : Word := 16#8371;   // error pending at kinematics
      ERR_MC_POWER : Word := 16#8372;   // error during execution of MC_POWER for axis
   END_VAR
   // statAxes[1].typeOfAxis := -1;
   // diagnostics.status := 16#7000;
   // startMode[1] := 1;
   // startMode[2] := 1;
   // startMode[3] := 1;
   // startMode[4] := 1;
BEGIN
   //==========================================================================================
   // SIEMENS AG
   // (c)Copyright 2020 All Rights Reserved
   //------------------------------------------------------------------------------------------
   // Library: LKinCtrl
   // Tested with: S7-1517T-3 PN/DP
   // Engineering: TIA Portal V15
   // Restrictions: ---
   // Requirements: S7-1500T FW 2.5
   // Functionality: LKinCtrl_MC_GroupPower
   // The FB is executing MC_RESET function blocks to reset all axes
   // and the axesGroup (TO Kinematics)
   // 
   // Support: tech.team.motioncontrol@siemens.com
   // Note: Parameter comments are only available in language 'English (United States)'
   //------------------------------------------------------------------------------------------
   // Change log table:
   // Version    Date          Expert in charge    Changes applied
   // 01.00.00   05.03.2019    JR                  First release version v1.0
   // 01.00.01   13.02.2020    FR                  Reset "axesEnabled" output in case of error
   //===========================================================================================

   #tempEnable := #enable; // Work with temporary value / create process image

   REGION ENABLING/DISABLING
     IF (#tempEnable = TRUE) AND (#statStatus = #STATUS_NO_CALL) THEN // Enable FB
       // First call; initialize FB
       #statBusy := TRUE;
       #statError := FALSE;
       #statAxesEnabled := FALSE;
       #statErrorUserCleared := FALSE;
       #statErrorAutoCleared := FALSE;
       #statStatus := #STATUS_FIRST_CALL;


       #statStateMachine := #DETECT_AXES; // State machine - start processing

       // initialize functionality: reset of variables, diagnostics, etc.
       #statDisablingCompleted := FALSE;
       #statAxisStatusWord := 16#0;
       #statExsitingAxesCtr := 0;
       #statDisabledAxesCtr := 0;
       #statEnabledAxesCtr := 0;
       #statErrorDetailNumber := 0;
       #statAxisNumberDiag := 0;
       #statSubfunctionStatus := #STATUS_NO_ERROR;


     ELSIF (#tempEnable = FALSE) AND (#statEnableOld = TRUE) THEN // Disable FB 
       #statStateMachine := #DISABLING_AXES;

     ELSIF (#statStatus = #STATUS_FIRST_CALL) THEN // Set status identifier of subsequent call
       #statStatus := #STATUS_SUBSEQUENT_CALL;
     END_IF;

     // Edge detection 'enable' input
     #statEnableOld := #tempEnable;
   END_REGION ENABLING/DISABLING

   IF (#statStatus = #STATUS_NO_CALL) THEN
     // Nothing to do -> End here to reduce "system load"
     RETURN;
   END_IF;

   REGION STATE_MACHINE
     CASE #statStateMachine OF // State machine of FB
       #NO_PROCESSING: // No processing active (Note: this state must always be present and left empty)
         ;

       #DETECT_AXES: // Processing active
         REGION DETECT_AXES
           // check available & connected axes at TO_Kinematics
           // assign DB number of connected axis to DB_ANY type
           IF #axesGroup.KinematicsAxis.A1 <> 0 THEN
             #statAxes[1].axis := #axesGroup.KinematicsAxis.A1;
             #statExsitingAxesCtr += 1;
           END_IF;
           IF #axesGroup.KinematicsAxis.A2 <> 0 THEN
             #statAxes[2].axis := #axesGroup.KinematicsAxis.A2;
             #statExsitingAxesCtr += 1;
           END_IF;
           IF #axesGroup.KinematicsAxis.A3 <> 0 THEN
             #statAxes[3].axis := #axesGroup.KinematicsAxis.A3;
             #statExsitingAxesCtr += 1;
           END_IF;
           IF #axesGroup.KinematicsAxis.A4 <> 0 THEN
             #statAxes[4].axis := #axesGroup.KinematicsAxis.A4;
             #statExsitingAxesCtr += 1;
           END_IF;

           // detect type of axis once for later call of corresponding FCs
           FOR #tempAxisCtr := 1 TO #MAX_NO_OF_AXES DO
             // check for axes to be existing
             IF #statAxes[#tempAxisCtr].axis <> 0 THEN
               IF TypeOfDB(#statAxes[#tempAxisCtr].axis) = TO_PositioningAxis THEN
                 // set type of axis to PosAxis
                 #statAxes[#tempAxisCtr].typeOfAxis := #TYPE_POSITIONING_AXIS;
               ELSIF TypeOfDB(#statAxes[#tempAxisCtr].axis) = TO_SynchronousAxis THEN
                 // set type of axis to PosAxis
                 #statAxes[#tempAxisCtr].typeOfAxis := #TYPE_SYNCHRONOUS_AXIS;
               END_IF;
             ELSE
               // set type of axis to 'not used'
               #statAxes[#tempAxisCtr].typeOfAxis := #AXIS_NOT_USED;
             END_IF;

           END_FOR;


           // go to next state
           #statStateMachine := #CHECK_AXES;
         END_REGION DETECT_AXES 

       #CHECK_AXES:
         REGION CHECK_AXES
           FOR #tempAxisCtr := 1 TO #MAX_NO_OF_AXES DO
             // check for axes to be existing
             IF #statAxes[#tempAxisCtr].typeOfAxis <> #AXIS_NOT_USED THEN
               // check type of axes used
               IF #statAxes[#tempAxisCtr].typeOfAxis = #TYPE_POSITIONING_AXIS THEN
                 // read TO_PositioningAxis status word
                 "LKinCtrl_GetPosAxisData"(posAxis := #statAxes[#tempAxisCtr].axis,
                                           statusWord => #statAxisStatusWord,
                                           errorDetailNumber => #statAxisErrorDetailNumber);
               ELSIF #statAxes[#tempAxisCtr].typeOfAxis = #TYPE_SYNCHRONOUS_AXIS THEN
                 // read TO_SynchronousAxis status word
                 "LKinCtrl_GetSyncAxisData"(syncAxis := #statAxes[#tempAxisCtr].axis,
                                            statusWord => #statAxisStatusWord,
                                            errorDetailNumber => #statAxisErrorDetailNumber);
               END_IF;
             END_IF;

             IF #statAxisStatusWord.%X1 = FALSE THEN
               // do nothing here, continue checks
               ;
             ELSE
               // set status
               #statStatus := #ERR_AXIS_ERROR;
               // set error bit
               #statErrorAutoCleared := TRUE;
               // write axis number to diagnostics
               #statAxisNumberDiag := #tempAxisCtr;
               // set subFunctionStatus
               #statErrorDetailNumber := #statAxisErrorDetailNumber;
               // go to error state
               #statStateMachine := #ERROR_STATE;
               EXIT;
             END_IF;

           END_FOR;

           // check TO_Kinematics to have no errors pending
           IF #axesGroup.StatusWord.%X1 = FALSE THEN
             // do nothing here, continue checks
             ;
           ELSE
             // check for no axis error detected prior
             IF #statAxisStatusWord.%X1 = FALSE THEN
               // set status
               #statStatus := #ERR_KIN_ERROR;
               // set error bit
               #statErrorAutoCleared := TRUE;
               // set subFunctionStatus
               #statErrorDetailNumber := #axesGroup.ErrorDetail.Number;
               // go to error state
               #statStateMachine := #ERROR_STATE;
             END_IF;

           END_IF;


           // check for no error to be pending
           IF #statStatus.%X15 = FALSE
             // // check MC_Power FBs to be not enabling the axes yet
             // AND #instMC_Power[1].Status = FALSE
             // AND #instMC_Power[2].Status = FALSE
             // AND #instMC_Power[3].Status = FALSE
             // AND #instMC_Power[4].Status = FALSE
           THEN
             // go to next state
             #statStateMachine := #ENABLING_AXES;
           END_IF;
         END_REGION CHECK_AXES

       #ENABLING_AXES: // Enabling active
         REGION ENABLING_AXES
           // set status message
           #statStatus := #STATUS_ENABLING_AXES_IN_PROGRESS;

           FOR #tempAxisCtr := 1 TO #MAX_NO_OF_AXES DO
             // check for axes to be existing
             IF #statAxes[#tempAxisCtr].typeOfAxis <> #AXIS_NOT_USED THEN
               // set execute trigger for MC_POWER
               #statEnableAxis[#tempAxisCtr] := TRUE;
             END_IF;
           END_FOR;


           // reset enabled axes counter
           #statEnabledAxesCtr := 0;
           // check for enabling to have completed successfully
           FOR #tempAxisCtr := 1 TO #MAX_NO_OF_AXES DO
             // only run code for existing axes
             IF #statAxes[#tempAxisCtr].typeOfAxis <> #AXIS_NOT_USED THEN
               // check for enabling to be done
               IF #instMC_Power[#tempAxisCtr].Status THEN
                 // count done signals
                 #statEnabledAxesCtr += 1;
               ELSIF #instMC_Power[#tempAxisCtr].Error THEN
                 // set status
                 #statStatus := #ERR_MC_POWER;
                 // set error bit
                 #statErrorAutoCleared := TRUE;
                 // write MC_HOME errorID to diagnostics
                 #statSubfunctionStatus := #instMC_Power[#tempAxisCtr].ErrorId;
                 // write axis number to diagnostics
                 #statAxisNumberDiag := #tempAxisCtr;
                 // exit FOR loop once error is found
                 EXIT;
                 // go to error state
                 #statStateMachine := #ERROR_STATE;
               END_IF;
             END_IF;
           END_FOR;

           // check for all axes to be enabled successfully
           IF #statEnabledAxesCtr = #statExsitingAxesCtr THEN
             // go to next state
             #statStateMachine := #ENABLED_AXES;
           END_IF;
         END_REGION ENABLING_AXES

       #ENABLED_AXES:
         REGION ENABLED_AXES
           // set output to signalize enabling successful
           #statAxesEnabled := TRUE;
           // set status message
           #statStatus := #STATUS_ALL_AXES_ENABLED;